      Appearance <- "DOx_DB_DD_CMD_Start_M"
   Button "Button_25" at 360,187 size 46x20; TextOff 'Inv'
      on Click: InvertBit("DOx_DB_DD_CMD_Inverse")
      Appearance <- "DOx_DB_DD_CMD_Inverse"
   Button "Button_26" at 360,212 size 46x20; TextOff 'Sim'
      on Click: InvertBit("DOx_DB_DD_CMD_Simulation")
      Appearance <- "DOx_DB_DD_CMD_Simulation"
   TextField "Text field_9" at 131,247 size 45x22; Text 'Q 0.4'
   TextField "Text field_10" at 176,247 size 119x22; Text 'Вибратор Пуск'
   Circle "Circle_9" at 131,270 size 22x22
      Appearance <- "DOx_DB_Vibro_CMD_Start_A"
   Circle "Circle_10" at 154,270 size 22x22
      Appearance <- "DOx_DB_Vibro_CMD_Q"
   Button "Button_27" at 298,248 size 59x44; TextOff 'Авто'; TextList "Hand"
      on Click: InvertBit("DOx_DB_Vibro_CMD_Hand")
      Appearance <- "DOx_DB_Vibro_CMD_Hand"
      ProcessValue <- "DOx_DB_Vibro_CMD_Hand"
   Button "Button_28" at 240,270 size 49x22; TextOff 'Выкл'
      on Click: ResetBit("DOx_DB_Vibro_CMD_Start_M")
   Button "Button_29" at 184,270 size 47x22; TextOff 'Вкл'
      on Click: SetBit("DOx_DB_Vibro_CMD_Start_M")
      Appearance <- "DOx_DB_Vibro_CMD_Start_M"
   Button "Button_30" at 360,247 size 46x20; TextOff 'Inv'
      on Click: InvertBit("DOx_DB_Vibro_CMD_Inverse")
      Appearance <- "DOx_DB_Vibro_CMD_Inverse"
   Button "Button_31" at 360,272 size 46x20; TextOff 'Sim'
      on Click: InvertBit("DOx_DB_Vibro_CMD_Simulation")
      Appearance <- "DOx_DB_Vibro_CMD_Simulation"
   TextField "Text field_11" at 131,306 size 45x22; Text 'Q 0.5'
   TextField "Text field_12" at 176,306 size 116x22; Text 'Жид.доз.Пуск'
   Circle "Circle_11" at 131,329 size 22x22
      Appearance <- "DOx_DB_DL_CMD_Start_A"
   Circle "Circle_12" at 154,329 size 22x22
      Appearance <- "DOx_DB_DL_CMD_Q"
   Button "Button_32" at 298,307 size 59x44; TextOff 'Авто'; TextList "Hand"
      on Click: InvertBit("DOx_DB_DL_CMD_Hand")
      Appearance <- "DOx_DB_DL_CMD_Hand"
      ProcessValue <- "DOx_DB_DL_CMD_Hand"
   Button "Button_33" at 240,329 size 49x22; TextOff 'Выкл'
      on Click: ResetBit("DOx_DB_DL_CMD_Start_M")
   Button "Button_34" at 184,329 size 47x22; TextOff 'Вкл'
      on Click: SetBit("DOx_DB_DL_CMD_Start_M")
      Appearance <- "DOx_DB_DL_CMD_Start_M"
   Button "Button_35" at 360,306 size 46x20; TextOff 'Inv'
      on Click: InvertBit("DOx_DB_DL_CMD_Inverse")
      Appearance <- "DOx_DB_DL_CMD_Inverse"
   Button "Button_36" at 360,331 size 46x20; TextOff 'Sim'
      on Click: InvertBit("DOx_DB_DL_CMD_Simulation")
      Appearance <- "DOx_DB_DL_CMD_Simulation"
   TextField "Text field_13" at 131,365 size 45x22; Text 'Q 0.6'
   TextField "Text field_14" at 176,365 size 110x22; Text 'КС1 Открыть'
   Circle "Circle_13" at 131,388 size 22x22
      Appearance <- "DOx_DB_KC1_CMD_Start_A"
   Circle "Circle_14" at 154,388 size 22x22
      Appearance <- "DOx_DB_KC1_CMD_Q"
   Button "Button_37" at 298,366 size 59x44; TextOff 'Авто'; TextList "Hand"
      on Click: InvertBit("DOx_DB_KC1_CMD_Hand")
      Appearance <- "DOx_DB_KC1_CMD_Hand"
      ProcessValue <- "DOx_DB_KC1_CMD_Hand"
   Button "Button_38" at 240,388 size 49x22; TextOff 'Выкл'
      on Click: ResetBit("DOx_DB_KC1_CMD_Start_M")
   Button "Button_39" at 184,388 size 47x22; TextOff 'Вкл'
      on Click: SetBit("DOx_DB_KC1_CMD_Start_M")
      Appearance <- "DOx_DB_KC1_CMD_Start_M"
   Button "Button_40" at 360,365 size 46x20; TextOff 'Inv'
      on Click: InvertBit("DOx_DB_KC1_CMD_Inverse")
      Appearance <- "DOx_DB_KC1_CMD_Inverse"
   Button "Button_41" at 360,390 size 46x20; TextOff 'Sim'
      on Click: InvertBit("DOx_DB_KC1_CMD_Simulation")
      Appearance <- "DOx_DB_KC1_CMD_Simulation"
   TextField "Text field_15" at 131,425 size 45x22; Text 'Q 0.7'
   TextField "Text field_16" at 176,425 size 117x22; Text 'LED Сухой ход'
   Circle "Circle_15" at 131,448 size 22x22
      Appearance <- "DOx_DB_LED_Dry_Run_Start_A"
   Circle "Circle_16" at 154,448 size 22x22
      Appearance <- "DOx_DB_LED_Dry_Run_Q"
   Button "Button_42" at 298,426 size 59x44; TextOff 'Авто'; TextList "Hand"
      on Click: InvertBit("DOx_DB_LED_Dry_Run_Hand")
      Appearance <- "DOx_DB_LED_Dry_Run_Hand"
      ProcessValue <- "DOx_DB_LED_Dry_Run_Hand"
   Button "Button_43" at 240,448 size 49x22; TextOff 'Выкл'
      on Click: ResetBit("DOx_DB_LED_Dry_Run_Start_M")
   Button "Button_44" at 184,448 size 47x22; TextOff 'Вкл'
      on Click: SetBit("DOx_DB_LED_Dry_Run_Start_M")
      Appearance <- "DOx_DB_LED_Dry_Run_Start_M"
   Button "Button_45" at 360,425 size 46x20; TextOff 'Inv'
      on Click: InvertBit("DOx_DB_LED_Dry_Run_Inverse")
      Appearance <- "DOx_DB_LED_Dry_Run_Inverse"
   Button "Button_46" at 360,450 size 46x20; TextOff 'Sim'
      on Click: InvertBit("DOx_DB_LED_Dry_Run_Simulation")
      Appearance <- "DOx_DB_LED_Dry_Run_Simulation"
   TextField "Text field_17" at 437,10 size 45x22; Text 'Q 1.0'
   TextField "Text field_18" at 482,10 size 93x22; Text 'LED Авария'
   Circle "Circle_17" at 437,33 size 22x22
      Appearance <- "DOx_DB_LED_Alarm_Start_A"
   Circle "Circle_18" at 460,33 size 22x22
      Appearance <- "DOx_DB_LED_Alarm_Q"
   Button "Button_47" at 604,11 size 59x44; TextOff 'Авто'; TextList "Hand"
      on Click: InvertBit("DOx_DB_LED_Alarm_Hand")
      Appearance <- "DOx_DB_LED_Alarm_Hand"
      ProcessValue <- "DOx_DB_LED_Alarm_Hand"
   Button "Button_48" at 546,33 size 49x22; TextOff 'Выкл'
      on Click: ResetBit("DOx_DB_LED_Alarm_Start_M")
   Button "Button_49" at 490,33 size 47x22; TextOff 'Вкл'
      on Click: SetBit("DOx_DB_LED_Alarm_Start_M")
      Appearance <- "DOx_DB_LED_Alarm_Start_M"
   Button "Button_50" at 666,10 size 46x20; TextOff 'Inv'
      on Click: InvertBit("DOx_DB_LED_Alarm_Inverse")
      Appearance <- "DOx_DB_LED_Alarm_Inverse"
   Button "Button_51" at 666,35 size 46x20; TextOff 'Sim'
      on Click: InvertBit("DOx_DB_LED_Alarm_Simulation")
      Appearance <- "DOx_DB_LED_Alarm_Simulation"
   TextField "Text field_19" at 437,69 size 45x22; Text 'Q 1.1'
   TextField "Text field_20" at 482,69 size 84x22; Text 'LED Пусто'
   Circle "Circle_19" at 437,92 size 22x22
      Appearance <- "DOx_DB_LED_Empty_Start_A"
   Circle "Circle_20" at 460,92 size 22x22
      Appearance <- "DOx_DB_LED_Empty_Q"
   Button "Button_52" at 604,70 size 59x44; TextOff 'Авто'; TextList "Hand"
      on Click: InvertBit("DOx_DB_LED_Empty_Hand")
      Appearance <- "DOx_DB_LED_Empty_Hand"
      ProcessValue <- "DOx_DB_LED_Empty_Hand"
   Button "Button_53" at 546,92 size 49x22; TextOff 'Выкл'
      on Click: ResetBit("DOx_DB_LED_Empty_Start_M")
   Button "Button_54" at 490,92 size 47x22; TextOff 'Вкл'
      on Click: SetBit("DOx_DB_LED_Empty_Start_M")
      Appearance <- "DOx_DB_LED_Empty_Start_M"
   Button "Button_55" at 666,69 size 46x20; TextOff 'Inv'
      on Click: InvertBit("DOx_DB_LED_Empty_Inverse")
      Appearance <- "DOx_DB_LED_Empty_Inverse"
   Button "Button_56" at 666,94 size 46x20; TextOff 'Sim'
      on Click: InvertBit("DOx_DB_LED_Empty_Simulation")
      Appearance <- "DOx_DB_LED_Empty_Simulation"
*)

(* ===== HMI "HMI_RT_1" =====
system functions are stored by id; their names below are inferred from use

graphic list "ok": 0 'check_box_off'; 1 'check_box_on'

graphic list "Status": 0 'sys_x'; 1 'sys_check-mark'; 2 'z2use'; 3 'alarm_on'

ScreenModuleEditorView "HMI_AI_full_R" 640x480
   Rectangle "Rectangle_2" at 176,16 size 320x270
      Visibility <- "View.view_settings"
   TextField "Text field_2" at 9,22 size 67x22; Text 'Датчик:'
   TextField "Text field_4" at 94,22 size 38x22; Text 'Text'
   TextField "Text field_6" at 287,14 size 147x22; Text 'Масштабирование'
      Visibility <- "View.view_settings"
   TextField "Text field_7" at 201,37 size 43x22; Text 'вход'
      Visibility <- "View.view_settings"
   TextField "Text field_8" at 201,62 size 56x22; Text 'выход'
      Visibility <- "View.view_settings"
   IOField "I/O field_1" at 267,38 size 92x26; FormatPattern s99999.9
      Visibility <- "View.view_settings"
      ProcessValue <- "AIx.C_Min_abs"
   IOField "I/O field_2" at 267,60 size 92x26; FormatPattern s99999.9
      Visibility <- "View.view_settings"
      ProcessValue <- "AIx.C_Min_out"
   IOField "I/O field_3" at 377,37 size 92x26; FormatPattern s99999.9
      Visibility <- "View.view_settings"
      ProcessValue <- "AIx.C_Max_abs"
   IOField "I/O field_4" at 377,59 size 92x26; FormatPattern s99999.9
      Visibility <- "View.view_settings"
      ProcessValue <- "AIx.C_Max_out"
   TextField "Text field_9" at 200,92 size 101x22; Text 'Фильтрация'
      Visibility <- "View.view_settings"
   TextField "Text field_10" at 201,117 size 36x22; Text 'RTD'
      Visibility <- "View.view_settings"
   Button "Button_1" at 311,95 size 20x20; TextOff 'Text'; PictureList "ok"
      on Click: InvertBit("AIx.F_Use")
      Visibility <- "View.view_settings"
      ProcessValue <- "AIx.F_Use"
   Button "Button_2" at 311,117 size 20x20; TextOff 'Text'; PictureList "ok"
      on Click: InvertBit("AIx.RTD")
      Visibility <- "View.view_settings"
      ProcessValue <- "AIx.RTD"
   IOField "I/O field_5" at 338,92 size 65x25; FormatPattern 9.99
      Visibility <- "View.view_settings"
      ProcessValue <- "AIx.F_Coeff"
   IOField "I/O field_6" at 338,117 size 65x25; FormatPattern 9999
      Visibility <- "View.view_settings"
      ProcessValue <- "AIx.RTD_C"
   TextField "Text field_11" at 11,53 size 79x22; Text 'Поправка'
   IOField "I/O field_7" at 94,53 size 78x23; FormatPattern s99.99
      ProcessValue <- "AIx.Calibration"
   Button "Button_3" at 201,200 size 68x28; TextOff 'Use'
      on Click: InvertBit("AIx.Use")
      Visibility <- "View.view_settings"
      Appearance <- "AIx.Use"
   Button "Button_4" at 14,85 size 68x28; TextOff 'Hand'
      on Click: InvertBit("AIx.Hand")
      Appearance <- "AIx.Hand"
   IOField "I/O field_8" at 94,85 size 78x28; FormatPattern s999.99
      ProcessValue <- "AIx.Result"
   TextField "Text field_12" at 248,149 size 27x22; Text 'NC'
      Visibility <- "View.view_settings"
   TextField "Text field_13" at 249,169 size 25x22; Text 'SC'
      Visibility <- "View.view_settings"
   TextField "Text field_14" at 8,160 size 27x22; Text 'HH'
   TextField "Text field_15" at 14,180 size 16x22; Text 'H'
   TextField "Text field_16" at 15,200 size 14x22; Text 'L'
   TextField "Text field_17" at 10,221 size 23x22; Text 'LL'
   IOField "I/O field_9" at 404,92 size 65x25; FormatPattern 99
      Visibility <- "View.view_settings"
      ProcessValue <- "AIx.F_SP"
   Button "Button_5" at 308,200 size 68x28; TextOff 'Invers'
      on Click: InvertBit("AIx.Inverse")
      Visibility <- "View.view_settings"
      Appearance <- "AIx.Inverse"
   IOField "I/O field_10" at 418,200 size 55x28; FormatPattern FFFF
      Visibility <- "View.view_settings"
      ProcessValue <- "AIx.Alarm"
   IOField "I/O field_11" at 284,149 size 58x21; FormatPattern s99999
      Visibility <- "View.view_settings"
      ProcessValue <- "AIx.A_SP_NC"
      Appearance <- "AIx.A_NC"
   IOField "I/O field_12" at 284,169 size 58x21; FormatPattern 99999
      Visibility <- "View.view_settings"
      ProcessValue <- "AIx.A_SP_SC"
      Appearance <- "AIx.A_SC"
   IOField "I/O field_13" at 44,160 size 58x21; FormatPattern s999.9
      ProcessValue <- "AIx.A_SP_HH"
      Appearance <- "AIx.A_HH"
   IOField "I/O field_14" at 44,180 size 58x21; FormatPattern s999.9
      ProcessValue <- "AIx.A_SP_H"
      Appearance <- "AIx.A_H"
   IOField "I/O field_15" at 44,200 size 58x21; FormatPattern s999.9
      ProcessValue <- "AIx.A_SP_L"
      Appearance <- "AIx.A_L"
   IOField "I/O field_16" at 44,220 size 58x21; FormatPattern s999.9
      ProcessValue <- "AIx.A_SP_LL"
      Appearance <- "AIx.A_LL"
   IOField "I/O field_17" at 358,149 size 58x21; FormatPattern 999
      Visibility <- "View.view_settings"
      ProcessValue <- "AIx.A_T_NC_SP"
   IOField "I/O field_18" at 358,169 size 58x21; FormatPattern 999
      Visibility <- "View.view_settings"
      ProcessValue <- "AIx.A_T_SC_SP"
   IOField "I/O field_19" at 118,160 size 58x21; FormatPattern 999
      ProcessValue <- "AIx.A_T_HH_SP"
   IOField "I/O field_20" at 118,180 size 58x21; FormatPattern 999
      ProcessValue <- "AIx.A_T_H_SP"
   IOField "I/O field_21" at 118,200 size 58x21; FormatPattern 999
      ProcessValue <- "AIx.A_T_L_SP"
   IOField "I/O field_22" at 118,220 size 58x21; FormatPattern 999
      ProcessValue <- "AIx.A_T_LL_SP"
   IOField "I/O field_23" at 404,117 size 65x25; FormatPattern 99999
      Visibility <- "View.view_settings"
      ProcessValue <- "AIx.Signal"
   TextField "Text field_18" at 8,132 size 68x22; Text 'Уставка'
   TextField "Text field_19" at 81,118 size 95x40; Text 'Время реакции (с)'
   Button "Button_6" at 80,247 size 96x32; TextOff 'Настройки'
      on Click: SetBit("View.view_settings")
   Button "Button_7" at 193,247 size 285x32; TextOff 'Сохранить'
      on Click: ResetBit("View.view_settings")
      Visibility <- "View.view_settings"
   GraphicIOField "Graphic I/O field_1" at 5,242 size 40x40; PictureList "Status"
      ProcessValue <- "AIx.Status"
*)

(* ===== HMI "HMI_RT_1" =====
system functions are stored by id; their names below are inferred from use

graphic list "ok": 0 'check_box_off'; 1 'check_box_on'

graphic list "Status": 0 'sys_x'; 1 'sys_check-mark'; 2 'z2use'; 3 'alarm_on'

ScreenModuleEditorView "HMI_AI_full_R" 640x480
   Rectangle "Rectangle_2" at 216,26 size 280x237
      Visibility <- "View.view_settings"
   TextField "Text field_2" at 49,27 size 67x22; Text 'Датчик:'
   TextField "Text field_4" at 121,27 size 38x22; Text 'Text'
   TextField "Text field_7" at 229,30 size 43x22; Text 'вход'
      Visibility <- "View.view_settings"
   TextField "Text field_8" at 229,55 size 56x22; Text 'выход'
      Visibility <- "View.view_settings"
   IOField "I/O field_1" at 295,31 size 92x26; FormatPattern s99999.9
      Visibility <- "View.view_settings"
      ProcessValue <- "AIx.C_Min_abs"
   IOField "I/O field_2" at 295,53 size 92x26; FormatPattern s99999.9
      Visibility <- "View.view_settings"
      ProcessValue <- "AIx.C_Min_out"
   IOField "I/O field_3" at 394,30 size 92x26; FormatPattern s99999.9
      Visibility <- "View.view_settings"
      ProcessValue <- "AIx.C_Max_abs"
   IOField "I/O field_4" at 394,52 size 92x26; FormatPattern s99999.9
      Visibility <- "View.view_settings"
      ProcessValue <- "AIx.C_Max_out"
   TextField "Text field_9" at 228,80 size 101x22; Text 'Фильтрация'
      Visibility <- "View.view_settings"
   TextField "Text field_10" at 229,105 size 36x22; Text 'RTD'
      Visibility <- "View.view_settings"
   Button "Button_1" at 328,83 size 20x20; TextOff 'Text'; PictureList "ok"
      on Click: InvertBit("AIx.F_Use")
      Visibility <- "View.view_settings"
      ProcessValue <- "AIx.F_Use"
   Button "Button_2" at 328,105 size 20x20; TextOff 'Text'; PictureList "ok"
      on Click: InvertBit("AIx.RTD")
      Visibility <- "View.view_settings"
      ProcessValue <- "AIx.RTD"
   IOField "I/O field_5" at 355,80 size 65x25; FormatPattern 9.99
      Visibility <- "View.view_settings"
      ProcessValue <- "AIx.F_Coeff"
   IOField "I/O field_6" at 355,105 size 65x25; FormatPattern 9999
      Visibility <- "View.view_settings"
      ProcessValue <- "AIx.RTD_C"
   TextField "Text field_11" at 49,48 size 79x22; Text 'Поправка'
   IOField "I/O field_7" at 132,48 size 78x23; FormatPattern s99.99
      ProcessValue <- "AIx.Calibration"
   Button "Button_3" at 235,180 size 68x28; TextOff 'Use'
      on Click: InvertBit("AIx.Use")
      Visibility <- "View.view_settings"
      Appearance <- "AIx.Use"
   Button "Button_4" at 52,78 size 68x28; TextOff 'Hand'
      on Click: InvertBit("AIx.Hand")
      Appearance <- "AIx.Hand"
   IOField "I/O field_8" at 132,78 size 78x28; FormatPattern s999.99
      ProcessValue <- "AIx.Result"
   TextField "Text field_12" at 270,135 size 27x22; Text 'NC'
      Visibility <- "View.view_settings"
   TextField "Text field_13" at 271,155 size 25x22; Text 'SC'
      Visibility <- "View.view_settings"
   TextField "Text field_14" at 49,137 size 27x22; Text 'HH'
   TextField "Text field_15" at 55,157 size 16x22; Text 'H'
   TextField "Text field_16" at 56,177 size 14x22; Text 'L'
   TextField "Text field_17" at 51,198 size 23x22; Text 'LL'
   IOField "I/O field_9" at 421,80 size 65x25; FormatPattern 99
      Visibility <- "View.view_settings"
      ProcessValue <- "AIx.F_SP"
   Button "Button_5" at 342,180 size 68x28; TextOff 'Invers'
      on Click: InvertBit("AIx.Inverse")
      Visibility <- "View.view_settings"
      Appearance <- "AIx.Inverse"
   IOField "I/O field_10" at 433,180 size 55x28; FormatPattern FFFF
      Visibility <- "View.view_settings"
      ProcessValue <- "AIx.Alarm"
   IOField "I/O field_11" at 306,135 size 58x21; FormatPattern s99999
      Visibility <- "View.view_settings"
      ProcessValue <- "AIx.A_SP_NC"
      Appearance <- "AIx.A_NC"
   IOField "I/O field_12" at 306,155 size 58x21; FormatPattern 99999
      Visibility <- "View.view_settings"
      ProcessValue <- "AIx.A_SP_SC"
      Appearance <- "AIx.A_SC"
   IOField "I/O field_13" at 85,137 size 58x21; FormatPattern s999.9
      ProcessValue <- "AIx.A_SP_HH"
      Appearance <- "AIx.A_HH"
   IOField "I/O field_14" at 85,157 size 58x21; FormatPattern s999.9
      ProcessValue <- "AIx.A_SP_H"
      Appearance <- "AIx.A_H"
   IOField "I/O field_15" at 85,177 size 58x21; FormatPattern s999.9
      ProcessValue <- "AIx.A_SP_L"
      Appearance <- "AIx.A_L"
   IOField "I/O field_16" at 85,197 size 58x21; FormatPattern s999.9
      ProcessValue <- "AIx.A_SP_LL"
      Appearance <- "AIx.A_LL"
   IOField "I/O field_17" at 380,135 size 58x21; FormatPattern 999
      Visibility <- "View.view_settings"
      ProcessValue <- "AIx.A_T_NC_SP"
   IOField "I/O field_18" at 380,155 size 58x21; FormatPattern 999
      Visibility <- "View.view_settings"
      ProcessValue <- "AIx.A_T_SC_SP"
   IOField "I/O field_19" at 159,137 size 58x21; FormatPattern 999
      ProcessValue <- "AIx.A_T_HH_SP"
   IOField "I/O field_20" at 159,157 size 58x21; FormatPattern 999
      ProcessValue <- "AIx.A_T_H_SP"
   IOField "I/O field_21" at 159,177 size 58x21; FormatPattern 999
      ProcessValue <- "AIx.A_T_L_SP"
   IOField "I/O field_22" at 159,197 size 58x21; FormatPattern 999
      ProcessValue <- "AIx.A_T_LL_SP"
   IOField "I/O field_23" at 421,105 size 65x25; FormatPattern 99999
      Visibility <- "View.view_settings"
      ProcessValue <- "AIx.Signal"
   TextField "Text field_18" at 49,109 size 68x22; Text 'Уставка'
   TextField "Text field_19" at 138,109 size 79x22; Text 'Время (с)'
   Button "Button_6" at 121,224 size 96x32; TextOff 'Настройки'
      on Click: SetBit("View.view_settings")
   Button "Button_7" at 234,223 size 257x32; TextOff 'Сохранить'
      on Click: ResetBit("View.view_settings")
      Visibility <- "View.view_settings"
   GraphicIOField "Graphic I/O field_1" at 46,219 size 40x40; PictureList "Status"
      ProcessValue <- "AIx.Status"
*)

(* ===== HMI "HMI_RT_1" =====
system functions are stored by id; their names below are inferred from use

HMI tags "Default tag table"
   "View_All" : Bool, internal

text list "Hand": 0 'Авто'; 1 'Ручной'

graphic list "Graphic_list_1": 0 'sys_x'; 1 'sys_check-mark'

ScreenModuleEditorView "HMI_AI_small_up" 640x480
   IOField "I/O field_1" at 52,132 size 61x32; FormatPattern 999.9
      ProcessValue <- "AI.Result"
      Appearance <- "AI.Alarm"
   TextField "Text field_1" at 113,139 size 15x22; Text 'C'
   Line "Line_1" at 35,135 size 0x25
      Visibility <- "AI.Alarm"
   Line "Line_2" at 35,135 size 0x25
      Visibility <- "AI.Alarm"
   Line "Line_3" at 35,135 size 0x25
      Visibility <- "AI.Alarm"
   Line "Line_4" at 35,135 size 0x25
      Visibility <- "AI.Alarm"
   Rectangle "Rectangle_2" at 15,30 size 120x99
      Visibility <- "View.view_circle"
   Button "Button_3" at 21,76 size 102x27; TextOff 'Авто'; TextList "Hand"
      on Click: InvertBit("AI.Hand")
      Appearance <- "AI.Hand"
      Visibility <- "View.view_circle"
      ProcessValue <- "AI.Hand"
   TextField "Text field_2" at 20,105 size 109x22; Text 'Text'
      Visibility <- "View.view_circle"
   IOField "I/O field_2" at 22,38 size 101x32; FormatPattern 999.9
      Visibility <- "View.view_circle"
      ObjectEnable <- "AI.Hand"
      Appearance <- "AI.Hand"
      ProcessValue <- "AI.Result"
   GraphicView "Graphics View" at 101,122 size 24x24; Picture "z2use"
      Visibility <- "AI.Hand"
   Button "Button_1" at 11,129 size 124x37; TextOff 'Text'
      on Click: InvertBit("View.view_circle")
   GraphicIOField "Graphic I/O field_1" at 23,135 size 25x25; PictureList "Graphic_list_1"
      Visibility <- "AI.Alarm"
      ProcessValue <- "AI.Use"
   GraphicView "Graphic view_1" at 23,136 size 25x25; Picture "error"
      Visibility <- "AI.Alarm"
   TextField "Text field_3" at 20,105 size 109x22; Text 'Text'
      Visibility <- "All"
*)

(* ===== HMI "HMI_RT_1" =====
system functions are stored by id; their names below are inferred from use

HMI tags "Default tag table"
   "View_All" : Bool, internal

text list "Hand": 0 'Авто'; 1 'Ручной'

graphic list "Graphic_list_1": 0 'sys_x'; 1 'sys_check-mark'

ScreenModuleEditorView "HMI_AI_small_down" 640x480
   IOField "I/O field_1" at 52,132 size 61x32; FormatPattern 999.9
      ProcessValue <- "AI.Result"
      Appearance <- "AI.Alarm"
   TextField "Text field_1" at 113,139 size 15x22; Text 'C'
   Line "Line_1" at 35,135 size 0x25
      Visibility <- "AI.Alarm"
   Line "Line_2" at 35,135 size 0x25
      Visibility <- "AI.Alarm"
   Line "Line_3" at 35,135 size 0x25
      Visibility <- "AI.Alarm"
   Line "Line_4" at 35,135 size 0x25
      Visibility <- "AI.Alarm"
   Rectangle "Rectangle_2" at 15,164 size 120x99
      Visibility <- "View.view_circle"
   Button "Button_3" at 23,230 size 102x27; TextOff 'Авто'; TextList "Hand"
      on Click: InvertBit("AI.Hand")
      Appearance <- "AI.Hand"
      Visibility <- "View.view_circle"
      ProcessValue <- "AI.Hand"
   TextField "Text field_2" at 21,167 size 109x22; Text 'Text'
      Visibility <- "View.view_circle"
   IOField "I/O field_2" at 24,192 size 101x32; FormatPattern 999.9
      Visibility <- "View.view_circle"
      ObjectEnable <- "AI.Hand"
      Appearance <- "AI.Hand"
      ProcessValue <- "AI.Result"
   GraphicView "Graphics View" at 101,122 size 24x24; Picture "z2use"
      Visibility <- "AI.Hand"
   Button "Button_1" at 11,129 size 124x37; TextOff 'Text'
      on Click: InvertBit("View.view_circle")
   GraphicIOField "Graphic I/O field_1" at 23,135 size 25x25; PictureList "Graphic_list_1"
      Visibility <- "AI.Alarm"
      ProcessValue <- "AI.Use"
   GraphicView "Graphic view_1" at 23,136 size 25x25; Picture "error"
      Visibility <- "AI.Alarm"
   TextField "Text field_3" at 21,167 size 109x22; Text 'Text'
      Visibility <- "All"
*)

(* ===== HMI "HMI_RT_1" =====
system functions are stored by id; their names below are inferred from use

graphic list "ok": 0 'check_box_off'; 1 'check_box_on'

graphic list "Status": 0 'sys_x'; 1 'sys_check-mark'; 2 'z2use'; 3 'alarm_on'

ScreenModuleEditorView "HMI_AI_full_L" 640x480
   Rectangle "Rectangle_2" at 33,53 size 320x270
      Visibility <- "View.view_settings"
   TextField "Text field_2" at 351,59 size 67x22; Text 'Датчик:'
   TextField "Text field_4" at 436,59 size 38x22; Text 'Text'
   TextField "Text field_6" at 144,51 size 147x22; Text 'Масштабирование'
      Visibility <- "View.view_settings"
   TextField "Text field_7" at 58,74 size 43x22; Text 'вход'
      Visibility <- "View.view_settings"
   TextField "Text field_8" at 58,99 size 56x22; Text 'выход'
      Visibility <- "View.view_settings"
   IOField "I/O field_1" at 124,75 size 92x26; FormatPattern s99999.9
      Visibility <- "View.view_settings"
      ProcessValue <- "AIx.C_Min_abs"
   IOField "I/O field_2" at 124,97 size 92x26; FormatPattern s99999.9
      Visibility <- "View.view_settings"
      ProcessValue <- "AIx.C_Min_out"
   IOField "I/O field_3" at 234,74 size 92x26; FormatPattern s99999.9
      Visibility <- "View.view_settings"
      ProcessValue <- "AIx.C_Max_abs"
   IOField "I/O field_4" at 234,96 size 92x26; FormatPattern s99999.9
      Visibility <- "View.view_settings"
      ProcessValue <- "AIx.C_Max_out"
   TextField "Text field_9" at 57,129 size 101x22; Text 'Фильтрация'
      Visibility <- "View.view_settings"
   TextField "Text field_10" at 58,154 size 36x22; Text 'RTD'
      Visibility <- "View.view_settings"
   Button "Button_1" at 168,132 size 20x20; TextOff 'Text'; PictureList "ok"
      on Click: InvertBit("AIx.F_Use")
      Visibility <- "View.view_settings"
      ProcessValue <- "AIx.F_Use"
   Button "Button_2" at 168,154 size 20x20; TextOff 'Text'; PictureList "ok"
      on Click: InvertBit("AIx.RTD")
      Visibility <- "View.view_settings"
      ProcessValue <- "AIx.RTD"
   IOField "I/O field_5" at 195,129 size 65x25; FormatPattern 9.99
      Visibility <- "View.view_settings"
      ProcessValue <- "AIx.F_Coeff"
   IOField "I/O field_6" at 195,154 size 65x25; FormatPattern 9999
      Visibility <- "View.view_settings"
      ProcessValue <- "AIx.RTD_C"
   TextField "Text field_11" at 353,90 size 79x22; Text 'Поправка'
   IOField "I/O field_7" at 436,90 size 78x23; FormatPattern s99.99
      ProcessValue <- "AIx.Calibration"
   Button "Button_3" at 58,237 size 68x28; TextOff 'Use'
      on Click: InvertBit("AIx.Use")
      Visibility <- "View.view_settings"
      Appearance <- "AIx.Use"
   Button "Button_4" at 356,122 size 68x28; TextOff 'Hand'
      on Click: InvertBit("AIx.Hand")
      Appearance <- "AIx.Hand"
   IOField "I/O field_8" at 436,122 size 78x28; FormatPattern s999.99
      ProcessValue <- "AIx.Result"
   TextField "Text field_12" at 105,186 size 27x22; Text 'NC'
      Visibility <- "View.view_settings"
   TextField "Text field_13" at 106,206 size 25x22; Text 'SC'
      Visibility <- "View.view_settings"
   TextField "Text field_14" at 350,197 size 27x22; Text 'HH'
   TextField "Text field_15" at 356,217 size 16x22; Text 'H'
   TextField "Text field_16" at 357,237 size 14x22; Text 'L'
   TextField "Text field_17" at 352,258 size 23x22; Text 'LL'
   IOField "I/O field_9" at 261,129 size 65x25; FormatPattern 99
      Visibility <- "View.view_settings"
      ProcessValue <- "AIx.F_SP"
   Button "Button_5" at 165,237 size 68x28; TextOff 'Invers'
      on Click: InvertBit("AIx.Inverse")
      Visibility <- "View.view_settings"
      Appearance <- "AIx.Inverse"
   IOField "I/O field_10" at 275,237 size 55x28; FormatPattern FFFF
      Visibility <- "View.view_settings"
      ProcessValue <- "AIx.Alarm"
   IOField "I/O field_11" at 141,186 size 58x21; FormatPattern s99999
      Visibility <- "View.view_settings"
      ProcessValue <- "AIx.A_SP_NC"
      Appearance <- "AIx.A_NC"
   IOField "I/O field_12" at 141,206 size 58x21; FormatPattern 99999
      Visibility <- "View.view_settings"
      ProcessValue <- "AIx.A_SP_SC"
      Appearance <- "AIx.A_SC"
   IOField "I/O field_13" at 386,197 size 58x21; FormatPattern s999.9
      ProcessValue <- "AIx.A_SP_HH"
      Appearance <- "AIx.A_HH"
   IOField "I/O field_14" at 386,217 size 58x21; FormatPattern s999.9
      ProcessValue <- "AIx.A_SP_H"
      Appearance <- "AIx.A_H"
   IOField "I/O field_15" at 386,237 size 58x21; FormatPattern s999.9
      ProcessValue <- "AIx.A_SP_L"
      Appearance <- "AIx.A_L"
   IOField "I/O field_16" at 386,257 size 58x21; FormatPattern s999.9
      ProcessValue <- "AIx.A_SP_LL"
      Appearance <- "AIx.A_LL"
   IOField "I/O field_17" at 215,186 size 58x21; FormatPattern 999
      Visibility <- "View.view_settings"
      ProcessValue <- "AIx.A_T_NC_SP"
   IOField "I/O field_18" at 215,206 size 58x21; FormatPattern 999
      Visibility <- "View.view_settings"
      ProcessValue <- "AIx.A_T_SC_SP"
   IOField "I/O field_19" at 460,197 size 58x21; FormatPattern 999
      ProcessValue <- "AIx.A_T_HH_SP"
   IOField "I/O field_20" at 460,217 size 58x21; FormatPattern 999
      ProcessValue <- "AIx.A_T_H_SP"
   IOField "I/O field_21" at 460,237 size 58x21; FormatPattern 999
      ProcessValue <- "AIx.A_T_L_SP"
   IOField "I/O field_22" at 460,257 size 58x21; FormatPattern 999
      ProcessValue <- "AIx.A_T_LL_SP"
   IOField "I/O field_23" at 261,154 size 65x25; FormatPattern 99999
      Visibility <- "View.view_settings"
      ProcessValue <- "AIx.Signal"
   TextField "Text field_18" at 350,169 size 68x22; Text 'Уставка'
   TextField "Text field_19" at 423,155 size 95x40; Text 'Время реакции (с)'
   Button "Button_6" at 422,284 size 96x32; TextOff 'Настройки'
      on Click: SetBit("View.view_settings")
   Button "Button_7" at 50,284 size 285x32; TextOff 'Сохранить'
      on Click: ResetBit("View.view_settings")
      Visibility <- "View.view_settings"
   GraphicIOField "Graphic I/O field_1" at 347,279 size 40x40; PictureList "Status"
      ProcessValue <- "AIx.Status"
*)

(* ===== HMI "HMI_RT_1" =====
system functions are stored by id; their names below are inferred from use

text list "Mode": 0 'Не используется'; 1 'Автоматический'; 2 'Ручной'

graphic list "ok": 0 'check_box_off'; 1 'check_box_on'

ScreenModuleEditorView "HMI_AO_full" 640x480
   TextField "Text field_1" at 43,31 size 251x22; Text 'Настройка аналогового выхода'
   TextField "Text field_2" at 35,60 size 99x22; Text 'Устройство:'
   TextField "Text field_3" at 35,85 size 57x22; Text 'Адрес:'
   TextField "Text field_4" at 135,60 size 38x22; Text 'Text'
   TextField "Text field_5" at 134,85 size 38x22; Text 'Text'
   TextField "Text field_6" at 123,107 size 147x22; Text 'Масштабирование'
   TextField "Text field_7" at 37,130 size 43x22; Text 'вход'
   TextField "Text field_8" at 37,155 size 56x22; Text 'выход'
   IOField "I/O field_1" at 103,131 size 92x26; FormatPattern s99999.9
      ProcessValue <- "AOx.C_Min_abs"
   IOField "I/O field_2" at 103,153 size 92x26; FormatPattern s99999.9
      ProcessValue <- "AOx.C_Min_out"
   IOField "I/O field_3" at 199,130 size 92x26; FormatPattern s99999.9
      ProcessValue <- "AOx.C_Max_abs"
   IOField "I/O field_4" at 199,152 size 92x26; FormatPattern s99999.9
      ProcessValue <- "AOx.C_Max_out"
   Button "Button_3" at 41,236 size 68x28; TextOff 'Use'
      on Click: InvertBit("AOx.Use")
      Appearance <- "AOx.Use"
   Button "Button_4" at 120,236 size 68x28; TextOff 'Hand'
      on Click: InvertBit("AOx.Hand")
      Appearance <- "AOx.Hand"
   IOField "I/O field_8" at 201,271 size 80x28; FormatPattern 99999
      ProcessValue <- "AOx.Signal"
   TextField "Text field_12" at 36,182 size 32x22; Text 'Min'
   TextField "Text field_13" at 37,207 size 36x22; Text 'Max'
   Button "Button_5" at 41,271 size 68x28; TextOff 'Invers'
      on Click: InvertBit("AOx.Inverse")
      Appearance <- "AOx.Inverse"
   Button "Button_6" at 120,271 size 68x28; TextOff 'Reset'
      on Click: InvertBit("AOx.Reset")
      Appearance <- "AOx.Reset"
   IOField "I/O field_11" at 75,182 size 58x21
      ProcessValue <- "AOx.Min"
   IOField "I/O field_12" at 75,207 size 58x21
      ProcessValue <- "AOx.Max"
   IOField "I/O field_13" at 195,181 size 58x21
      ProcessValue <- "AOx.Step_up"
   IOField "I/O field_14" at 195,206 size 58x21
      ProcessValue <- "AOx.Step_down"
   IOField "I/O field_23" at 241,83 size 58x21; FormatPattern s999.9
      ProcessValue <- "AOx.SP"
   Button "Button_1" at 135,182 size 56x20; TextOff 'Up'
      on Click: InvertBit("AOx.Up_use")
      Appearance <- "AOx.Up_use"
   Button "Button_2" at 135,208 size 56x20; TextOff 'Down'
      on Click: InvertBit("AOx.Down_use")
      Appearance <- "AOx.Down_use"
   IOField "I/O field_5" at 201,236 size 80x28; FormatPattern 999.9
      ProcessValue <- "AOx.Hand_SP"
   IOField "I/O field_6" at 257,181 size 45x21; FormatPattern 99.9
      ProcessValue <- "AOx.T_Up_SP"
   IOField "I/O field_7" at 257,206 size 45x21; FormatPattern 99.9
      ProcessValue <- "AOx.T_Down_SP"
*)

(* ===== HMI "HMI_RT_1" =====
system functions are stored by id; their names below are inferred from use

text list "Mode": 0 'Не используется'; 1 'Автоматический'; 2 'Ручной'

graphic list "ok": 0 'check_box_off'; 1 'check_box_on'

ScreenModuleEditorView "HMI_AO_full" 640x480
   TextField "Text field_2" at 35,74 size 99x22; Text 'Устройство:'
   TextField "Text field_3" at 35,101 size 57x22; Text 'Адрес:'
   TextField "Text field_4" at 135,74 size 38x22; Text 'Text'
   TextField "Text field_5" at 134,101 size 38x22; Text 'Text'
   TextField "Text field_7" at 37,130 size 43x22; Text 'вход'
   TextField "Text field_8" at 37,155 size 56x22; Text 'выход'
   IOField "I/O field_1" at 103,131 size 92x26; FormatPattern s99999.9
      ProcessValue <- "AOx.C_Min_abs"
   IOField "I/O field_2" at 103,153 size 92x26; FormatPattern s99999.9
      ProcessValue <- "AOx.C_Min_out"
   IOField "I/O field_3" at 210,130 size 92x26; FormatPattern s99999.9
      ProcessValue <- "AOx.C_Max_abs"
   IOField "I/O field_4" at 210,152 size 92x26; FormatPattern s99999.9
      ProcessValue <- "AOx.C_Max_out"
   Button "Button_3" at 41,236 size 68x28; TextOff 'Use'
      on Click: InvertBit("AOx.Use")
      Appearance <- "AOx.Use"
   Button "Button_4" at 131,236 size 68x28; TextOff 'Hand'
      on Click: InvertBit("AOx.Hand")
      Appearance <- "AOx.Hand"
   IOField "I/O field_8" at 221,271 size 80x28; FormatPattern 99999
      ProcessValue <- "AOx.Signal"
   TextField "Text field_12" at 36,182 size 32x22; Text 'Min'
   TextField "Text field_13" at 37,207 size 36x22; Text 'Max'
   Button "Button_5" at 41,271 size 68x28; TextOff 'Invers'
      on Click: InvertBit("AOx.Inverse")
      Appearance <- "AOx.Inverse"
   Button "Button_6" at 131,271 size 68x28; TextOff 'Reset'
      on Click: InvertBit("AOx.Reset")
      Appearance <- "AOx.Reset"
   IOField "I/O field_11" at 75,182 size 58x21
      ProcessValue <- "AOx.Min"
   IOField "I/O field_12" at 75,207 size 58x21
      ProcessValue <- "AOx.Max"
   IOField "I/O field_13" at 195,181 size 58x21
      ProcessValue <- "AOx.Step_up"
   IOField "I/O field_14" at 195,206 size 58x21
      ProcessValue <- "AOx.Step_down"
   IOField "I/O field_23" at 243,103 size 58x21; FormatPattern s999.9
      ProcessValue <- "AOx.SP"
   Button "Button_1" at 135,182 size 56x20; TextOff 'Up'
      on Click: InvertBit("AOx.Up_use")
      Appearance <- "AOx.Up_use"
   Button "Button_2" at 135,208 size 56x20; TextOff 'Down'
      on Click: InvertBit("AOx.Down_use")
      Appearance <- "AOx.Down_use"
   IOField "I/O field_5" at 221,236 size 80x28; FormatPattern 999.9
      ProcessValue <- "AOx.Hand_SP"
   IOField "I/O field_6" at 257,181 size 45x21; FormatPattern 99.9
      ProcessValue <- "AOx.T_Up_SP"
   IOField "I/O field_7" at 257,206 size 45x21; FormatPattern 99.9
      ProcessValue <- "AOx.T_Down_SP"
*)

(* ===== HMI "HMI_RT_1" =====
system functions are stored by id; their names below are inferred from use

text list "Hand": 0 'Авто'; 1 'Ручной'

ScreenModuleEditorView "HMI_DI_full" 640x480
   TextField "Text field_1" at 16,21 size 34x22; Text 'I x.x'
   TextField "Text field_2" at 59,21 size 68x22; Text 'not used'
   Circle "Circle_1" at 16,44 size 22x22
      Appearance <- "DIx.Input"
   Circle "Circle_2" at 16,67 size 22x22
      Appearance <- "DIx.Start"
   Button "Button_3" at 43,45 size 95x20; TextOff 'Авто'; TextList "Hand"
      on Click: InvertBit("DIx.Hand")
      ProcessValue <- "DIx.Hand"
      Appearance <- "DIx.Hand"
   Button "Button_4" at 89,67 size 49x20; TextOff 'Выкл'
      on Click: ResetBit("DIx.Start")
   Button "Button_12" at 43,67 size 47x20; TextOff 'Вкл'
      on Click: SetBit("DIx.Start")
      Appearance <- "DIx.Start"
   TextField "Text field_16" at 139,49 size 29x18; Text 'Вкл:'
   IOField "I/O field_6" at 177,47 size 30x20; FormatPattern 99
      ProcessValue <- "DIx.ON_SP"
   IOField "I/O field_7" at 177,67 size 30x20; FormatPattern 99
      ProcessValue <- "DIx.OFF_SP"
   TextField "Text field_17" at 140,67 size 37x18; Text 'Выкл:'
   Button "Button_1" at 178,24 size 60x20; TextOff 'Inv'
      on Click: InvertBit("DIx.Inverse")
      Appearance <- "DIx.Inverse"
   IOField "I/O field_1" at 209,47 size 30x20; FormatPattern 99
      ProcessValue <- "DIx.ON_Now"
   IOField "I/O field_2" at 209,67 size 30x20; FormatPattern 99
      ProcessValue <- "DIx.OFF_Now"
*)

(* ===== HMI "HMI_RT_1" =====
system functions are stored by id; their names below are inferred from use

text list "Hand": 0 'Авто'; 1 'Ручной'

ScreenModuleEditorView "HMI_DO_full" 640x480
   TextField "Text field_1" at 16,21 size 38x22; Text 'Q x.x'
   TextField "Text field_2" at 65,21 size 68x22; Text 'not used'
   Circle "Circle_1" at 16,44 size 22x22
      Appearance <- "DOx.Signal"
   Circle "Circle_2" at 16,67 size 22x22
      Appearance <- "DOx.Output"
   Button "Button_3" at 43,45 size 95x20; TextOff 'Авто'; TextList "Hand"
      on Click: InvertBit("DOx.Hand")
      Appearance <- "DOx.Hand"
      ProcessValue <- "DOx.Hand"
   Button "Button_4" at 89,67 size 49x20; TextOff 'Выкл'
      on Click: ResetBit("DOx.Output")
   Button "Button_12" at 43,67 size 47x20; TextOff 'Вкл'
      on Click: SetBit("DOx.Output")
      Appearance <- "DOx.Output"
   Button "Button_1" at 148,45 size 60x20; TextOff 'Inv'
      on Click: InvertBit("DOx.Inverse")
      Appearance <- "DOx.Inverse"
   Button "Button_2" at 148,68 size 60x20; TextOff 'Sim'
      on Click: InvertBit("DOx.Simultation")
      Appearance <- "DOx.Simultation"
   Button "Button_5" at 148,21 size 60x20; TextOff 'Imp'
      on Click: InvertBit("DOx.Impulse")
      Appearance <- "DOx.Impulse"
   IOField "I/O field_6" at 214,45 size 30x20; FormatPattern 99
      Visibility <- "DOx.Impulse"
      ProcessValue <- "DOx.T_SP"
   IOField "I/O field_7" at 214,68 size 30x20; FormatPattern 99
      Visibility <- "DOx.Impulse"
      ProcessValue <- "DOx.T_Now"
   TextField "Text field_3" at 212,26 size 40x15; Text '100ms'
      Visibility <- "DOx.Impulse"
*)

(* ===== HMI "HMI_RT_1" =====
system functions are stored by id; their names below are inferred from use

text list "Number": 1 'P1'; 2 'P2'; 3 'P3'; 4 'P11-A'; 5 'P12-A'; 6 'P13-A'; 7 'P14-I'; 8 'P15'; 9 'P4'; 10 'P6-A'; 11 'P7-A'; 12 'P21-A'; 13 'P22-A'; 14 'P10'; 15 'P11'; 16 'P12'; 17 'IE-P-02'; 18 'P26-I'; 19 'P27'; 20 'S27'; 21 'P24'; 22 'P25-A'; 23 'P25'; 24 'P29-A'; 25 'P31-A'; 26 'P33'; 27 'P25'; 28 'P26'; 29 'DP11'; 30 'DP12'; 31 'DP23'; 32 'DP65'

text list "Mode": 0 'Автомат'; 1 'Ручной'; 2 'Force'; 3 'Симуляция'; 4 'Удалённый'; 5 'Локальный'; 6 'Заблокирован'; 7 ''; 8 ''; 9 'Отключён'; 10 'Сервисный'

text list "Status": 0 'Выкл'; 1 'Вкл'; 2 'Остановка'; 3 'Запуск'; 4 'Авария ВЫКЛ'; 5 'Авария ВКЛ'; 6 'Авария QF'; 7 'Отключён'

text list "Hand": 0 'Авто'; 1 'Ручной'

graphic list "Start_M": 0 'off'; 1 'on_2'

graphic list "Pump_Down": 1 'pump_ok'; 2 'pump_wait'; 3 'pump_wait_1'; 7 'down_stop'; 0 'pump_off'; 4 'pump'; 8 'down_start'; 9 'down_alm'

graphic list "Pump_Left": 1 'left_on'; 2 'left_wait'; 3 'left_wait_1'; 7 'left_stop'; 0 'left_off'; 4 'left_no'; 8 'left_start'; 9 'left_alm'

graphic list "Pump_Right": 1 'right_on'; 2 'right_wait'; 3 'right_wait_1'; 7 'right_stop'; 0 'right_off'; 4 'right_no'; 8 'right_start'; 9 'right_alm'

graphic list "Pump_Up": 1 'up_on'; 2 'up_wait'; 3 'up_wait'; 7 'up_stop'; 0 'up_off'; 4 'up_no'; 8 'up_start'; 9 'up_alm'

graphic list "V_Down": 1 'down_open_3x'; 2 'down_closing_3x'; 3 'down_opening_3x'; 7 'down_cl_alm_3xя'; 0 'down_close_3x'; 4 'down_no_3x'; 8 'down_op_alm_3x'; 9..100 'down_alm_3x'

graphic list "V_Left": 1 'left_open_3x'; 2 'left_closing_3x'; 3 'left_opening_3x'; 7 'left_cl_alm_3xя'; 0 'left_close_3x'; 4 'left_no_3x'; 8 'left_op_alm_3x'; 9..100 'left_alm_3x'

graphic list "V_Right": 1 'right_open_3x'; 2 'right_closing_3x'; 3 'right_opening_3x'; 7 'right_cl_alm_3xя'; 0 'right_close_3x'; 4 'right_no_3x'; 8 'right_op_alm_3x'; 9..100 'right_alm_3x'

graphic list "V_Up": 1 'up_open_3x'; 2 'up_closing_3x'; 3 'up_opening_3x'; 7 'up_cl_alm_3xя'; 0 'up_close_3x'; 4 'up_no_3x'; 8 'up_op_alm_3x'; 9 'up_alm_3x'

graphic list "Z_Hor": 1 'h_open'; 2 'd_closing'; 3 'd_opening_1'; 0 'v_close'; 4 'v_no'; 7..100 'down_alm_3x'

graphic list "Z_Vert": 1 'v_open'; 2 'd_closing_1'; 3 'd_opening'; 0 'h_close'; 4 'h_no'; 7..100 'h_alarm'

ScreenModuleEditorView "HMI_M_Uni_DA_micro" 1024x768
   Button "Button_2" at 100,82 size 41x40; TextOff 'Text'; PictureList "Start_M"
      on Click: InvertBit("Motor.Start_M")
      Visibility <- "Visu.view_circle"
      ObjectEnable <- "Motor.Hand"
      ProcessValue <- "Motor.Start_M"
   Circle "Circle_7" at 137,109 size 47x47
      Visibility <- "Motor.Sim"
   GraphicIOField "Graphic I/O field_1" at 146,118 size 30x30; PictureList "Pump_Down"
      Visibility <- "Type"
      ProcessValue <- "Motor.Status"
   GraphicView "Graphic view_11" at 119,101 size 30x30; Picture "service"
      Visibility <- "Motor.Trace_lock"
   GraphicIOField "Graphic I/O field_2" at 146,118 size 30x30; PictureList "Pump_Up"
      Visibility <- "Type"
      ProcessValue <- "Motor.Status"
   GraphicIOField "Graphic I/O field_3" at 146,118 size 30x30; PictureList "Pump_Left"
      Visibility <- "Type"
      ProcessValue <- "Motor.Status"
   GraphicIOField "Graphic I/O field_4" at 146,118 size 30x30; PictureList "Pump_Right"
      Visibility <- "Type"
      ProcessValue <- "Motor.Status"
   IOField "I/O field_1" at 134,149 size 55x30; FormatPattern 999.9
      Visibility <- "Motor.Analog"
      ObjectEnable <- "Motor.Hand"
      Appearance <- "Motor.Hand"
      ProcessValue <- "Motor.SP_M"
   GraphicView "Graphic view_8" at 170,134 size 30x30; Picture "force"
      Visibility <- "Motor.Force"
   GraphicView "Graphic view_12" at 121,132 size 30x30; Picture "local"
      Visibility <- "Motor.Local"
   GraphicView "Graphic view_4" at 185,125 size 38x37; Picture "z2_2"
      Visibility <- "Visu.view_circle"
   Button "Button_5" at 184,122 size 43x44; TextOff 'Text'
      on Click: ResetBit("Motor.Hand"); ResetBit("Visu.view_settings"); ResetBit("Visu.view_alm"); ResetBit("Visu.view_circle")
      Visibility <- "Visu.view_circle"
      ObjectEnable <- "Visu.view_circle"
   GraphicView "Graphic view_6" at 103,122 size 38x37; Picture "z2_1"
      Visibility <- "Visu.view_circle"
   Button "Button_6" at 102,117 size 39x44; TextOff 'Text'
      on Click: SetBit("Motor.Hand"); ResetBit("Visu.view_settings"); ResetBit("Visu.view_alm"); ResetBit("Visu.view_circle")
      Visibility <- "Visu.view_circle"
      ObjectEnable <- "Visu.view_circle"
   GraphicIOField "Graphic I/O field_5" at 146,118 size 30x30; PictureList "V_Down"
      Visibility <- "Type"
      ProcessValue <- "Motor.Status"
   GraphicIOField "Graphic I/O field_6" at 146,118 size 30x30; PictureList "V_Up"
      Visibility <- "Type"
      ProcessValue <- "Motor.Status"
   GraphicIOField "Graphic I/O field_7" at 146,118 size 30x30; PictureList "V_Left"
      Visibility <- "Type"
      ProcessValue <- "Motor.Status"
   GraphicIOField "Graphic I/O field_8" at 146,118 size 30x30; PictureList "V_Right"
      Visibility <- "Type"
      ProcessValue <- "Motor.Status"
   GraphicIOField "Graphic I/O field_9" at 146,118 size 30x30; PictureList "Z_Hor"
      Visibility <- "Type"
      ProcessValue <- "Motor.Status"
   GraphicIOField "Graphic I/O field_10" at 146,118 size 30x30; PictureList "Z_Vert"
      Visibility <- "Type"
      ProcessValue <- "Motor.Status"
   GraphicView "Graphic view_10" at 146,117 size 30x30; Picture "lock_32x32"
      Visibility <- "Motor.Lock"
   Button "Button_13" at 137,109 size 48x51; TextOff 'Text'
      on Click: InvertBit("Visu.view_circle"); ResetBit("Visu.view_alm"); ResetBit("Visu.view_settings")
   IOField "I/O field_3" at 136,85 size 55x30; FormatPattern 999.9
      Visibility <- "Motor.Analog"
      ProcessValue <- "Motor.FB_SP"
   TextField "Text field_13" at 121,79 size 85x26; Text 'Text'
      Visibility <- "Visu.view_circle"
   TextField "Text field_1" at 121,79 size 85x26; Text 'Text'
      Visibility <- "All"
   GraphicView "Graphic view_7" at 174,101 size 30x30; Picture "z2_1"
      Visibility <- "Motor.Hand"
*)

(* ===== HMI "HMI_RT_1" =====
system functions are stored by id; their names below are inferred from use

text list "Mode": 0 'ПИ'; 1 'ПИД'

graphic list "ok": 0 'check_box_off'; 1 'check_box_on'

ScreenModuleEditorView "HMI_PID_ex" 640x480
   TextField "Text field_7" at 292,39 size 43x22; Text 'вход'
      Visibility <- "Visu.view_settings"
   TextField "Text field_8" at 292,64 size 56x22; Text 'выход'
      Visibility <- "Visu.view_settings"
   IOField "I/O field_1" at 358,40 size 92x26; FormatPattern s99999.9
      Visibility <- "Visu.view_settings"
      ProcessValue <- "PIDx.Min_in"
   IOField "I/O field_2" at 358,62 size 92x26; FormatPattern s99999.9
      Visibility <- "Visu.view_settings"
      ProcessValue <- "PIDx.Min_out"
   IOField "I/O field_3" at 454,39 size 92x26; FormatPattern s99999.9
      Visibility <- "Visu.view_settings"
      ProcessValue <- "PIDx.Max_in"
   IOField "I/O field_4" at 454,61 size 92x26; FormatPattern s99999.9
      Visibility <- "Visu.view_settings"
      ProcessValue <- "PIDx.Max_out"
   Button "Button_6" at 290,115 size 68x30; TextOff 'Reset'
      on Click: SetBit("PIDx.Reset")
      Visibility <- "Visu.view_settings"
      Appearance <- "PIDx.Reset"
   IOField "I/O field_10" at 360,115 size 55x30; FormatPattern FFFF
      Visibility <- "Visu.view_settings"
      ProcessValue <- "PIDx.Warning_code"
   TextField "Text field_5" at 288,152 size 46x22; Text 'Cycle'
      Visibility <- "Visu.view_settings"
   IOField "I/O field_9" at 343,152 size 63x23; FormatPattern 99.9
      Visibility <- "Visu.view_settings"
      ProcessValue <- "PIDx.SP_Cycle"
   IOField "I/O field_15" at 417,115 size 55x30; FormatPattern FFFF
      Visibility <- "Visu.view_settings"
      ProcessValue <- "PIDx.Error_code"
      Appearance <- "PIDx.Error"
   Button "Button_2" at 475,115 size 71x30; TextOff 'Invers'
      on Click: InvertBit("PIDx.Invert")
      Visibility <- "Visu.view_settings"
      Appearance <- "PIDx.Invert"
   TextField "Text field_17" at 292,87 size 67x22; Text 'уставка'
      Visibility <- "Visu.view_settings"
   IOField "I/O field_17" at 358,85 size 92x26; FormatPattern s99999.9
      Visibility <- "Visu.view_settings"
      ProcessValue <- "PIDx.Min_out"
   IOField "I/O field_18" at 454,84 size 92x26; FormatPattern s99999.9
      Visibility <- "Visu.view_settings"
      ProcessValue <- "PIDx.Max_out"
   TextField "Text field_14" at 415,150 size 62x22; Text 'OnTime'
      Visibility <- "Visu.view_settings"
   IOField "I/O field_13" at 480,150 size 63x23; FormatPattern 99.9
      Visibility <- "Visu.view_settings"
      ProcessValue <- "PIDx.OnTime"
   TextField "Text field_15" at 416,180 size 65x22; Text 'OffTime'
      Visibility <- "Visu.view_settings"
   IOField "I/O field_14" at 481,180 size 63x23; FormatPattern 99.9
      Visibility <- "Visu.view_settings"
      ProcessValue <- "PIDx.OffTime"
   TextField "Text field_18" at 288,208 size 102x22; Text 'SP Low Limit'
      Visibility <- "Visu.view_settings"
      Appearance <- "PIDx.SP_L"
   TextField "Text field_19" at 438,208 size 105x22; Text 'SP High Limit'
      Visibility <- "Visu.view_settings"
      Appearance <- "PIDx.SP_H"
   TextField "Text field_20" at 288,232 size 98x22; Text 'In Low Limit'
      Visibility <- "Visu.view_settings"
      Appearance <- "PIDx.In_L"
   TextField "Text field_21" at 438,232 size 101x22; Text 'In High Limit'
      Visibility <- "Visu.view_settings"
      Appearance <- "PIDx.In_H"
   Rectangle "Rectangle_2" at 237,26 size 320x268
      Visibility <- "Visu.view_settings"
   TextField "Text field_1" at 45,31 size 219x22; Text 'Настройка ПИД регулятора'
   TextField "Text field_2" at 35,60 size 101x22; Text 'Назначение:'
   TextField "Text field_4" at 136,61 size 38x22; Text 'Text'
   TextField "Text field_9" at 38,115 size 15x22; Text 'K'
   TextField "Text field_10" at 38,147 size 19x22; Text 'Ti'
   IOField "I/O field_5" at 76,117 size 70x30; FormatPattern s999.99
      ProcessValue <- "PIDx.SP_P"
   IOField "I/O field_6" at 76,148 size 70x30; FormatPattern 999.9
      ProcessValue <- "PIDx.SP_Ti"
   TextField "Text field_11" at 38,180 size 23x22; Text 'Td'
   IOField "I/O field_7" at 76,179 size 70x30; FormatPattern 999.9
      ProcessValue <- "PIDx.SP_Td"
   Button "Button_4" at 78,220 size 68x30; TextOff 'Hand'
      on Click: InvertBit("PIDx.Hand")
      Appearance <- "PIDx.Hand"
   IOField "I/O field_8" at 41,257 size 109x30; FormatPattern s999.99
      ProcessValue <- "PIDx.HandValue"
   SymbolicIOField "Symbolic I/O field_1" at 103,83 size 81x24; TextOn '1'; TextOff '0'; TextList "Mode"
      ProcessValue <- "PIDx.Type"
   TextField "Text field_3" at 34,81 size 62x22; Text 'Режим:'
   TextField "Text field_12" at 182,115 size 67x22; Text 'Датчик:'
   IOField "I/O field_11" at 181,137 size 63x23; FormatPattern s999.9
      ProcessValue <- "PIDx.Value"
   TextField "Text field_13" at 176,177 size 73x22; Text 'Уставка:'
   IOField "I/O field_12" at 182,201 size 63x23; FormatPattern s999.9
      ProcessValue <- "PIDx.SP"
   IOField "I/O field_16" at 176,260 size 77x28; FormatPattern s999.9
      ProcessValue <- "PIDx.Result"
   TextField "Text field_16" at 186,238 size 53x22; Text 'Result'
   Button "Button_1" at 40,220 size 30x30; TextOff 'Text'; PictureOff "sys_volume control"
      on Click: SetBit("Visu.view_settings")
   Button "Button_3" at 287,259 size 255x30; TextOff 'Save'
      on Click: ResetBit("Visu.view_settings")
      Visibility <- "Visu.view_settings"
*)

(* ===== HMI "HMI_RT_1" =====
system functions are stored by id; their names below are inferred from use

text list "Mode": 0 'ПИ'; 1 'ПИД'

graphic list "ok": 0 'check_box_off'; 1 'check_box_on'

